// TIA Portal project "Energy_Drink_V15.1" (V15.1) (continued)

       // IF RESET BUTTON OR HMI RESET => RESET RECIPE SELCTION
       IF "Reset_Button" OR "HMI_VAR".Reset_Selection THEN
           "RECIPE_1_DB".Recipe1.Recipe_Act := FALSE;
           "RECIPE_2_DB".Recipe2.Recipe_Act := FALSE;
           "RECIPE_3_DB".Recipe3.Recipe_Act := FALSE;
           "TEST_RECIPE_DB".Test.Recipe_Act := FALSE;
           "Recipe_Num" := 0;
       END_IF;

   END_REGION

   (************************ RECIPE CONFIRMARTION MANAGEMENT **********************************)
   REGION RECIPE SELECTION CONFIRMATION

       // IF ENTER SELECTION IS PRESSED => START PROCESS
       IF "Var_System_DB".System_Generic.Enter_Selection THEN
           "Var_System_DB".System_Generic.Man_Start_Process := true;
       END_IF;

       // IF ENTER SELECTION IS PRESSED => START PROCESS
       IF "HMI_VAR".Enter_Selection THEN
           "HMI_VAR".Start_Process := TRUE;
       END_IF;

   END_REGION
END_FUNCTION

// folder: 05-CONVEYOR MANAGEMENT

FUNCTION "CONVEYOR_BELT" : Void   // FC10, FBD
{ S7_Optimized_Access := 'FALSE' }
VERSION : 0.1
   VAR_INPUT
      Conveyor_Cmd : Bool;
      Time_Act : Time;
   END_VAR
BEGIN

REGION Network 1 (STL): *******************COMMANDS AND CONDITIONS TO MANAGE CONVEYOR BELT********************************************/
   // WHEN SCALE IS FINISHED WEIGHING ALL THE PRODUCTS => BACH IN PROGRESS =1
   // SEND COMMAND TO ACTIVATE THE CONVEYOR BELT
         A     #Conveyor_Cmd;
         FP    "FP_Conveyor_Act";
         S     "Var_System_DB".System_Generic.Mixer_Station;

         A     "Var_System_DB".System_Generic.Mixer_Station;
         FP    "Tag_14";
         =     "Var_System_DB".Conveyor_Belt.Motor_Cmd;


   // TIMER ACTIVATION: IF FN PULSE OF CONVEYOR_CMD => SET TIMER_ACT
         A     #Conveyor_Cmd;
         FN    "FN_Bach_in_Prog";
         =     "Var_System_DB".Conveyor_Belt.Timer_Act;

   // IF TIMER_ACT = 1 => ACTIVATE TIMER
         CALL  TP, "T_CONVEYOR"
         ( IN := "Var_System_DB".Conveyor_Belt.Timer_Act,
           PT := #Time_Act,
           Q  := ,
           ET :=
         );


   // IF TIMER.Q => SEND PULSE TO RESET MOTOR_CMD
         A     "T_CONVEYOR".Q;
         FN    "FN_TIMER.Q";
         R     "Var_System_DB".Conveyor_Belt.M_Stop;


   // SEND PULSE TO SET STOP COMMAND TO ITS NORMAL POSITON "NC" WHEN FN OF FEEDBACK
         A     "Var_System_DB".Conveyor_Belt.M_Feedback;
         FN    "FN_STOP_CMD";
         S     "Var_System_DB".Conveyor_Belt.M_Stop;
         S     "Var_System_DB".System_Generic.Conveyor_Station;


   // RESET CONVEYOR STATION
         A     "AGITATOR_TIMER_DB".Q;
         R     "Var_System_DB".System_Generic.Conveyor_Station;

   // MOTOR MEMORY STATE: IN CASE STOP BUTTON IS PRESSED AND THE  MOTOR WAS ACTIVE,
   // WE WANT TO KEEP THE MOTOR "ON" AFTER THE STOP BUTTON IS REALESED AGAIN
         A     "Var_System_DB".Conveyor_Belt.M_Feedback;
         S     "Var_System_DB".Conveyor_Belt.State;

   // RESET BELT STATE BIT
         AN    "Var_System_DB".System_Generic.Stop_Process;
         AN    "Var_System_DB".System_Generic.System_Failure;
         O(;
         A     "Var_System_DB".System_Generic.Start;
         FN    "Tag_27";
         );
         R     "Var_System_DB".Conveyor_Belt.State;
END_REGION

REGION Network 2: ****************** CONVEYOR BELT MOTOR ACTIVATION********************************************/
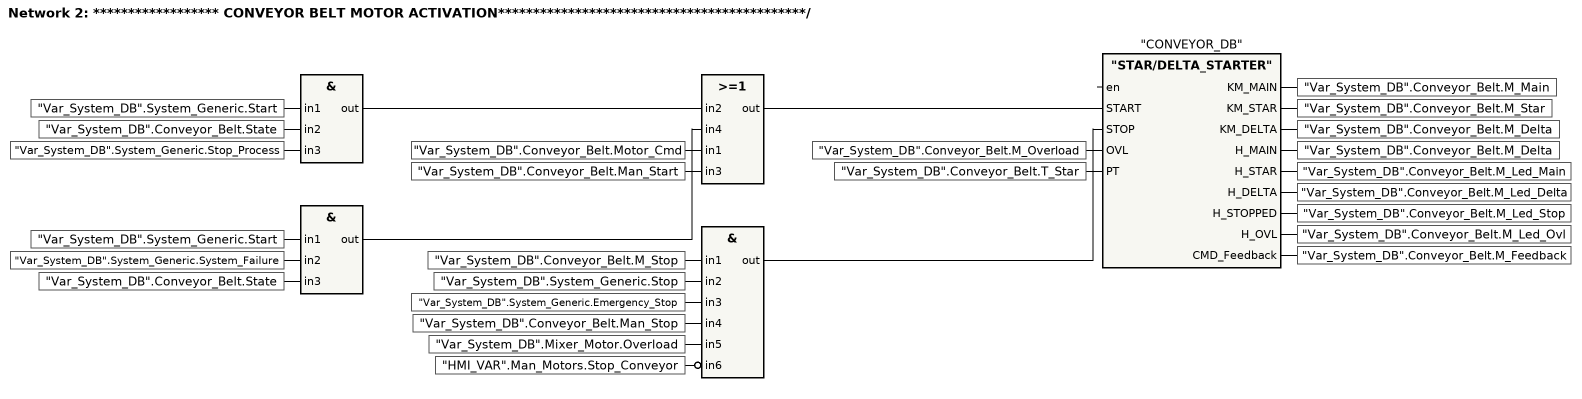
   "CONVEYOR_DB"(START := ("Var_System_DB".System_Generic.Start AND "Var_System_DB".Conveyor_Belt.State AND "Var_System_DB".System_Generic.Stop_Process) OR ("Var_System_DB".System_Generic.Start AND "Var_System_DB".System_Generic.System_Failure AND "Var_System_DB".Conveyor_Belt.State) OR "Var_System_DB".Conveyor_Belt.Motor_Cmd OR "Var_System_DB".Conveyor_Belt.Man_Start,   // "STAR/DELTA_STARTER"
                 STOP := "Var_System_DB".Conveyor_Belt.M_Stop AND "Var_System_DB".System_Generic.Stop AND "Var_System_DB".System_Generic.Emergency_Stop AND "Var_System_DB".Conveyor_Belt.Man_Stop AND "Var_System_DB".Mixer_Motor.Overload AND NOT "HMI_VAR".Man_Motors.Stop_Conveyor,
                 OVL := "Var_System_DB".Conveyor_Belt.M_Overload,
                 PT := "Var_System_DB".Conveyor_Belt.T_Star,
                 KM_MAIN => "Var_System_DB".Conveyor_Belt.M_Main,
                 KM_STAR => "Var_System_DB".Conveyor_Belt.M_Star,
                 KM_DELTA => "Var_System_DB".Conveyor_Belt.M_Delta,
                 H_MAIN => "Var_System_DB".Conveyor_Belt.M_Delta,
                 H_STAR => "Var_System_DB".Conveyor_Belt.M_Led_Main,
                 H_DELTA => "Var_System_DB".Conveyor_Belt.M_Led_Delta,
                 H_STOPPED => "Var_System_DB".Conveyor_Belt.M_Led_Stop,
                 H_OVL => "Var_System_DB".Conveyor_Belt.M_Led_Ovl,
                 CMD_Feedback => "Var_System_DB".Conveyor_Belt.M_Feedback);
END_REGION
END_FUNCTION

// folder: 06-MIXER MANAGEMENT

FUNCTION "MIXER_TANK_MANAGEMENT" : Void   // FC3, FBD
{ S7_Optimized_Access := 'FALSE' }
VERSION : 0.1
BEGIN

REGION Network 1: /***********************MIXER TANK LEVEL*****************************************/
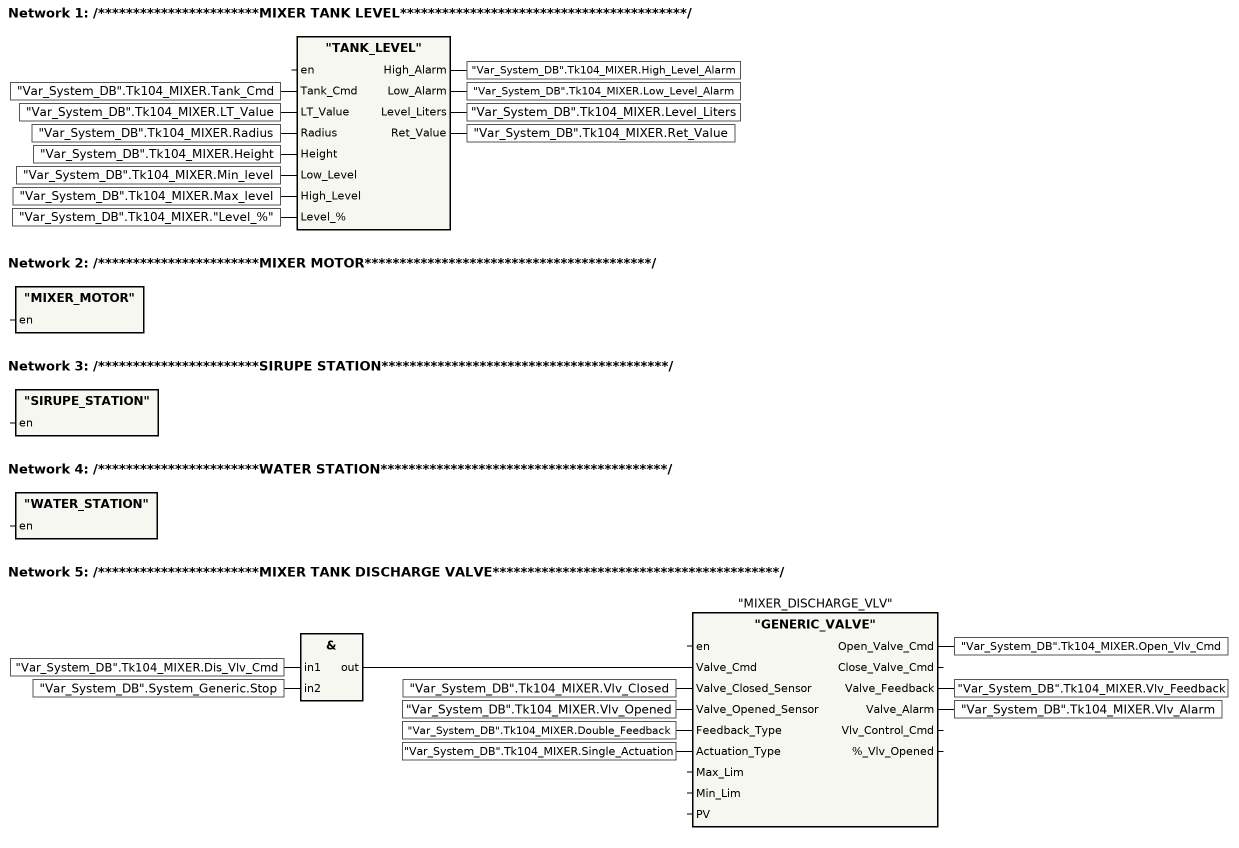
   "TANK_LEVEL"(Tank_Cmd := "Var_System_DB".Tk104_MIXER.Tank_Cmd,
                LT_Value := "Var_System_DB".Tk104_MIXER.LT_Value,
                Radius := "Var_System_DB".Tk104_MIXER.Radius,
                Height := "Var_System_DB".Tk104_MIXER.Height,
                Low_Level := "Var_System_DB".Tk104_MIXER.Min_level,
                High_Level := "Var_System_DB".Tk104_MIXER.Max_level,
                "Level_%" := "Var_System_DB".Tk104_MIXER."Level_%",
                High_Alarm => "Var_System_DB".Tk104_MIXER.High_Level_Alarm,
                Low_Alarm => "Var_System_DB".Tk104_MIXER.Low_Level_Alarm,
                Level_Liters => "Var_System_DB".Tk104_MIXER.Level_Liters,
                Ret_Value => "Var_System_DB".Tk104_MIXER.Ret_Value);
END_REGION

REGION Network 2: /***********************MIXER MOTOR*****************************************/
   "MIXER_MOTOR"();
END_REGION

REGION Network 3: /***********************SIRUPE STATION*****************************************/
   "SIRUPE_STATION"();
END_REGION

REGION Network 4: /***********************WATER STATION*****************************************/
   "WATER_STATION"();
END_REGION

REGION Network 5: /***********************MIXER TANK DISCHARGE VALVE*****************************************/
   "MIXER_DISCHARGE_VLV"(Valve_Cmd := "Var_System_DB".Tk104_MIXER.Dis_Vlv_Cmd AND "Var_System_DB".System_Generic.Stop,   // "GENERIC_VALVE"
                         Valve_Closed_Sensor := "Var_System_DB".Tk104_MIXER.Vlv_Closed,
                         Valve_Opened_Sensor := "Var_System_DB".Tk104_MIXER.Vlv_Opened,
                         Feedback_Type := "Var_System_DB".Tk104_MIXER.Double_Feedback,
                         Actuation_Type := "Var_System_DB".Tk104_MIXER.Single_Actuation,
                         Open_Valve_Cmd => "Var_System_DB".Tk104_MIXER.Open_Vlv_Cmd,
                         Valve_Feedback => "Var_System_DB".Tk104_MIXER.Vlv_Feedback,
                         Valve_Alarm => "Var_System_DB".Tk104_MIXER.Vlv_Alarm);
END_REGION

REGION Network 6 (STL): /***********************TANK CONDITIONS ACTIVATION*****************************************/
   // IF SYSTEM IS ACTIVE AND MIXER STATION => MIXER TANK COMMAND = 1
         A     "Var_System_DB".System_Generic.System_Act;
         A     "Var_System_DB".System_Generic.Mixer_Station;
         =     "Var_System_DB".Tk104_MIXER.Tank_Cmd;

   // IF TANK LEVEL > 15% => SEND COMMAND TO AGITATOR, WATER AND SIRUPE VALVE
         A     "Var_System_DB".Tk104_MIXER.Tank_Cmd;
         A(;
         L     "Var_System_DB".Tk104_MIXER."Level_%";
         L     15;
         >I;
         );
         =     "Var_System_DB".Mixer_Motor.Motor_Cmd;
         =     "Var_System_DB".Sirupe_Valve.Vlv_Cmd;
         =     "Var_System_DB".Water_Valve.Vlv_Cmd;
END_REGION

REGION Network 7 (STL): /***********************TANK CONDITIONS ACTIVATION*****************************************/
   // IF SYSTEM IS ACTIVE, MIXER STATION AND CONVEYOR HAS STOPPED =>
   // ACTIVATE TIMER TO OPEN THE VALVE WHEN ELAPSED TIME IS "ON"
         A     "Var_System_DB".System_Generic.System_Act;
         A     "Var_System_DB".System_Generic.Mixer_Station;
         A     "Var_System_DB".System_Generic.Conveyor_Station;
         FP    "Var_System_DB".Mixer_Motor.FP_Timer;
         =     "Var_System_DB".System_Generic.T_Mixer_Station;

   // TIMER CALL
         CALL  TP, "AGITATOR_TIMER_DB"
         ( IN := "Var_System_DB".System_Generic.T_Mixer_Station,
           PT := T#60S,
           Q  := ,
           ET :=
         );


   // IF FN AGITATOR_TIMER.Q => SEND COMMAND TO ACTIVATE DISCHARGE VALVE
         A     "AGITATOR_TIMER_DB".Q;
         FN    "Var_System_DB".Tk104_MIXER.FN_Agitator;
         S     "Var_System_DB".Tk104_MIXER.Dis_Vlv_Cmd;


   // RESET VALVE COMMAND AND MIXER STATION AND BACH IN PROGRESS
         A     "Var_System_DB".Tk104_MIXER.Dis_Vlv_Cmd;
         A(;
         L     "Var_System_DB".Tk104_MIXER."Level_%";
         L     0;
         ==I;
         );
         R     "Var_System_DB".Tk104_MIXER.Dis_Vlv_Cmd;
         R     "Var_System_DB".System_Generic.Mixer_Station;
         R     "Var_System_DB".System_Generic.Bach_In_Progress;

         ON    "Var_System_DB".System_Generic.System_Act;
         R     "Var_System_DB".Tk104_MIXER.Dis_Vlv_Cmd;
END_REGION
END_FUNCTION

FUNCTION "WATER_STATION" : Void   // FC5, FBD
{ S7_Optimized_Access := 'FALSE' }
VERSION : 0.1
BEGIN

REGION Network 1 (STL): /************************WATER FLOW METER*****************************************/
         CALL  SCALE
         ( IN      := "Var_System_DB".Water_Flow_Meter.Flow_Meter,
           HI_LIM  := "Var_System_DB".Water_Flow_Meter.High_Lim,
           LO_LIM  := "Var_System_DB".Water_Flow_Meter.Low_Lim,
           BIPOLAR := FALSE,
           RET_VAL := "Var_System_DB".Water_Flow_Meter.Ret_Val,
           OUT     := "Var_System_DB".Water_Flow_Meter.Flow_PV
         );
END_REGION

REGION Network 2: /*****************************WATER VALVE***************************************************/
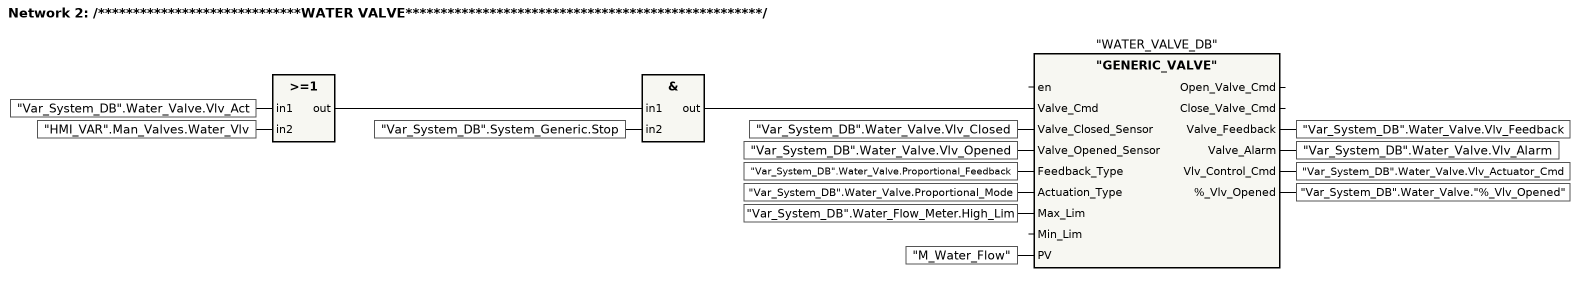
   "WATER_VALVE_DB"(Valve_Cmd := ("Var_System_DB".Water_Valve.Vlv_Act OR "HMI_VAR".Man_Valves.Water_Vlv) AND "Var_System_DB".System_Generic.Stop,   // "GENERIC_VALVE"
                    Valve_Closed_Sensor := "Var_System_DB".Water_Valve.Vlv_Closed,
                    Valve_Opened_Sensor := "Var_System_DB".Water_Valve.Vlv_Opened,
                    Feedback_Type := "Var_System_DB".Water_Valve.Proportional_Feedback,
                    Actuation_Type := "Var_System_DB".Water_Valve.Proportional_Mode,
                    Max_Lim := "Var_System_DB".Water_Flow_Meter.High_Lim,
                    PV := "M_Water_Flow",
                    Valve_Feedback => "Var_System_DB".Water_Valve.Vlv_Feedback,
                    Valve_Alarm => "Var_System_DB".Water_Valve.Vlv_Alarm,
                    Vlv_Control_Cmd => "Var_System_DB".Water_Valve.Vlv_Actuator_Cmd,
                    "%_Vlv_Opened" => "Var_System_DB".Water_Valve."%_Vlv_Opened");
END_REGION

REGION Network 3 (STL)
   // IF VALVE COMMAND SEND PULSE TO ACTIVATE => WATER VALVE
         A     "Var_System_DB".Water_Valve.Vlv_Cmd;
         FP    "Var_System_DB".Water_Valve.FP_Start;
         S     "Var_System_DB".Water_Valve.Vlv_Act;

   // IF MIXWE DISCHARGE VALVE COMMAND SEND PULSE TO DEACTIVATE => WATER VALVE
         A     "Var_System_DB".Tk104_MIXER.Dis_Vlv_Cmd;
         FP    "Var_System_DB".Water_Valve.FP_Stop;
         R     "Var_System_DB".Water_Valve.Vlv_Act;
END_REGION
END_FUNCTION

FUNCTION "SIRUPE_STATION" : Void   // FC7, FBD
{ S7_Optimized_Access := 'FALSE' }
VERSION : 0.1
BEGIN

REGION Network 1 (STL): /************************SIRUPE FLOW METER*****************************************/
         CALL  SCALE
         ( IN      := "Var_System_DB".Sirupe_Flow_Meter.Flow_Meter,
           HI_LIM  := "Var_System_DB".Sirupe_Flow_Meter.Low_Lim,
           LO_LIM  := "Var_System_DB".Sirupe_Flow_Meter.High_Lim,
           BIPOLAR := FALSE,
           RET_VAL := "Var_System_DB".Sirupe_Flow_Meter.Ret_Val,
           OUT     := "Var_System_DB".Sirupe_Flow_Meter.Flow_PV
         );
END_REGION

REGION Network 2 (STL)
         L     "M_Sirupe_Flow";
         L     1000;
         *R;
         T     "Var_System_DB".Sirupe_Valve.Increment_T;
END_REGION

REGION Network 3: /**********************************SIRUPE VALVE*****************************************/
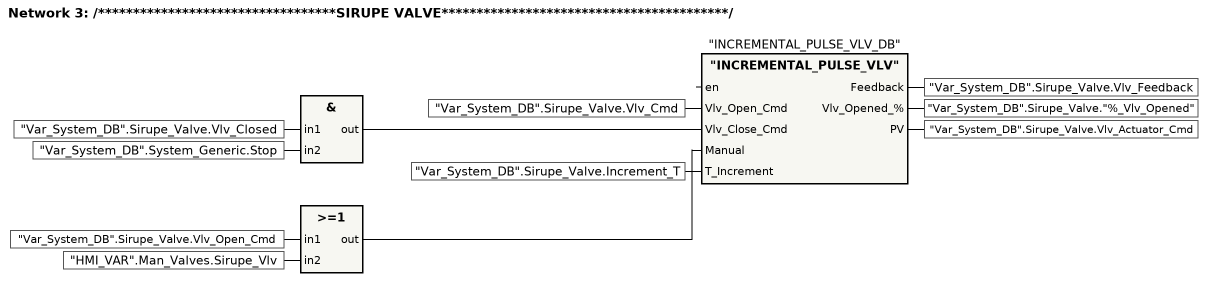
   "INCREMENTAL_PULSE_VLV_DB"(Vlv_Open_Cmd := "Var_System_DB".Sirupe_Valve.Vlv_Cmd,   // "INCREMENTAL_PULSE_VLV"
                           Vlv_Close_Cmd := "Var_System_DB".Sirupe_Valve.Vlv_Closed AND "Var_System_DB".System_Generic.Stop,
                           Manual := "Var_System_DB".Sirupe_Valve.Vlv_Open_Cmd OR "HMI_VAR".Man_Valves.Sirupe_Vlv,
                           T_Increment := "Var_System_DB".Sirupe_Valve.Increment_T,
                           Feedback => "Var_System_DB".Sirupe_Valve.Vlv_Feedback,
                           "Vlv_Opened_%" => "Var_System_DB".Sirupe_Valve."%_Vlv_Opened",
                           PV => "Var_System_DB".Sirupe_Valve.Vlv_Actuator_Cmd);
END_REGION

REGION Network 4 (STL)
   // COMMAND TO CLOSE THE VALVE
         A     "Var_System_DB".Tk104_MIXER.Dis_Vlv_Cmd;
         FP    "Var_System_DB".Sirupe_Valve.FP_Reset;
         =     "Var_System_DB".Sirupe_Valve.Vlv_Closed;
END_REGION
END_FUNCTION

FUNCTION "MIXER_MOTOR" : Void   // FC13, FBD
{ S7_Optimized_Access := 'FALSE' }
VERSION : 0.1
BEGIN

REGION Network 1 (STL): *******************COMMANDS AND CONDITIONS TO MANAGE AGITATOR********************************************/
   // IF MOTOR CMD FP => SEND COMMAND TO ACTIVATE AGITATOR
         A     "Var_System_DB".Mixer_Motor.Motor_Cmd;
         FP    "Var_System_DB".Mixer_Motor.FP_Start;
         O     "Var_System_DB".Mixer_Motor.Man_Start;
         =     "Var_System_DB".Mixer_Motor.Cmd_Start;

   // IF MOTOR CMD FN => SEND COMMAND TO DEACTIVATE AGITATOR
         A     "Var_System_DB".Mixer_Motor.Motor_Cmd;
         FN    "Var_System_DB".Mixer_Motor.FN_Stop;
         ON    "Var_System_DB".Mixer_Motor.Man_Stop;
         R     "Var_System_DB".Mixer_Motor.Cmd_Stop;


   // IF CMD STOP NOT ACTIVE AND MOTOR PV = 0 => SET BACK CMD STOP = 1
         AN    "Var_System_DB".Mixer_Motor.Cmd_Stop;
         A(;
         L     "Var_System_DB".Mixer_Motor.PV;
         L     0;
         ==I;
         );
         S     "Var_System_DB".Mixer_Motor.Cmd_Stop;


   // RESET MIXER MOTOR STATE:
   // IF NOT STOP PROCESS AND NOT SYSTEM FAILURE (NOT OVERLOAD) AND MOTOR_PV == 0
   // OR NEGATIVE EDGE OF GENERIC START
         AN    "Var_System_DB".System_Generic.Stop_Process;
         AN    "Var_System_DB".System_Generic.System_Failure;
         A(;
         L     "Var_System_DB".Mixer_Motor.PV;
         L     0;
         ==I;
         );
         O(;
         A     "Var_System_DB".System_Generic.Start;
         FN    "Tag_26";
         );
         R     "Var_System_DB".Mixer_Motor.State;


   // MOTOR MEMORY STATE IN CASE STOP BUTTON PRESSED AND THE  MOTOR WAS ACTIVE
   // WE WANT TO KEEP THE MOTOR ON AFTER THE STOP BUTTON
         A     "Var_System_DB".Mixer_Motor.Feedback;
         S     "Var_System_DB".Mixer_Motor.State;
END_REGION

REGION Network 2
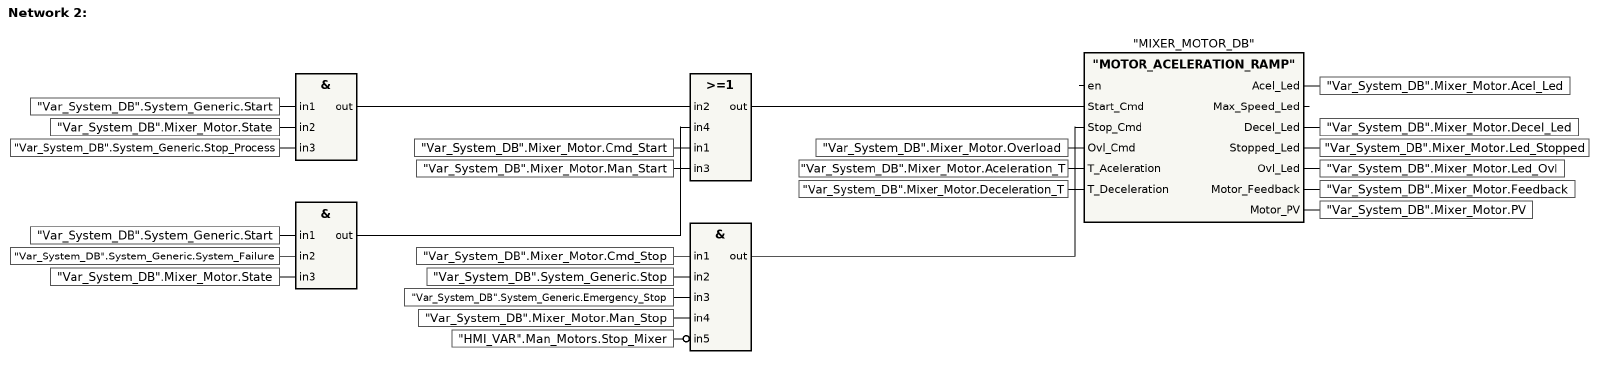
   "MIXER_MOTOR_DB"(Start_Cmd := ("Var_System_DB".System_Generic.Start AND "Var_System_DB".Mixer_Motor.State AND "Var_System_DB".System_Generic.Stop_Process) OR ("Var_System_DB".System_Generic.Start AND "Var_System_DB".System_Generic.System_Failure AND "Var_System_DB".Mixer_Motor.State) OR "Var_System_DB".Mixer_Motor.Cmd_Start OR "Var_System_DB".Mixer_Motor.Man_Start,   // "MOTOR_ACELERATION_RAMP"
                    Stop_Cmd := "Var_System_DB".Mixer_Motor.Cmd_Stop AND "Var_System_DB".System_Generic.Stop AND "Var_System_DB".System_Generic.Emergency_Stop AND "Var_System_DB".Mixer_Motor.Man_Stop AND NOT "HMI_VAR".Man_Motors.Stop_Mixer,
                    Ovl_Cmd := "Var_System_DB".Mixer_Motor.Overload,
                    T_Aceleration := "Var_System_DB".Mixer_Motor.Aceleration_T,
                    T_Deceleration := "Var_System_DB".Mixer_Motor.Deceleration_T,
                    Acel_Led => "Var_System_DB".Mixer_Motor.Acel_Led,
                    Decel_Led => "Var_System_DB".Mixer_Motor.Decel_Led,
                    Stopped_Led => "Var_System_DB".Mixer_Motor.Led_Stopped,
                    Ovl_Led => "Var_System_DB".Mixer_Motor.Led_Ovl,
                    Motor_Feedback => "Var_System_DB".Mixer_Motor.Feedback,
                    Motor_PV => "Var_System_DB".Mixer_Motor.PV);
END_REGION
END_FUNCTION

// folder: FBs

FUNCTION_BLOCK "GENERIC_VALVE"   // FB1, SCL
{ S7_Optimized_Access := 'FALSE' }
VERSION : 0.1
   VAR_INPUT
      Valve_Cmd : Bool;   // Enable valve command
      Valve_Closed_Sensor : Bool;   // Valve closed position
      Valve_Opened_Sensor : Bool;   // Valve opened position
      Feedback_Type : Int;   // "0" = No feedback / "1"= Single disFeedback / "2"= Single EnFeedback / "3" = Double Feedback / "4" = Proportional
      Actuation_Type : Int;
      Max_Lim : Real;
      Min_Lim : Real;
      PV : Real;
   END_VAR
   VAR_OUTPUT
      Open_Valve_Cmd : Bool;
      Close_Valve_Cmd : Bool;
      Valve_Feedback : Bool;   // "1" If the valve is open, "0" otherwise
      Valve_Alarm : Bool;
      Vlv_Control_Cmd : Int;
      "%_Vlv_Opened" : DInt;
   END_VAR
   VAR
      M_Vlv_Closed : Bool;
      M_Vlv_Opened : Bool;
      Ret_Vlv : Word;
   END_VAR
   VAR_TEMP
      Temp_Process_Signal : Real;
   END_VAR
   VAR CONSTANT
      No_Feedback : Int := 0;
      Single_En_Feedback : Int := 1;
      Single_Dis_Feedback : Int := 2;
      Double_Feedback : Int := 3;
      Proportional_Feedback : Int := 4;
      Single_Actuation : Int := 1;
      Double_Actuation : Int := 2;
      Proportional_Mode : Int := 3;
      Inverse_Mode : Int := 4;
      Control_Loop : Int := 5;
   END_VAR
BEGIN
   (*
   *File: FB GENERIC VALVE 
   * Author: Jaime Calvente Mieres
   * Date: 18-05-2022
   * Description: This FB will be used to control a valve. Depending on 
     the users input, the valve could act as Single actuation,
     Double actuation or Proportional mode.
   *)



   (*This Case Statement will be used to map the process sensors to
   the internal variables used for the program logic, based on the
   Feedback Type or (Type of Valve) used in each process.*)
   REGION FEEDBACK_TYPE

       CASE #Feedback_Type OF

           #No_Feedback:
               ;

           #Single_En_Feedback:
               #M_Vlv_Opened := #Valve_Opened_Sensor;

           #Single_Dis_Feedback:
               #M_Vlv_Closed := #Valve_Closed_Sensor;

           #Double_Feedback:
               #M_Vlv_Closed := #Valve_Closed_Sensor;
               #M_Vlv_Opened := #Valve_Opened_Sensor;

           #Proportional_Feedback:
               #M_Vlv_Closed := #Valve_Closed_Sensor;
               #M_Vlv_Opened := #Valve_Opened_Sensor;

           ELSE  // Statement section ELSE
               ;
       END_CASE;


   END_REGION


   // IF VALVE COMMAND ACTIVE
   IF #Valve_Cmd THEN

   (*This Case Statement will be used to Set the type of Actuation will be used
   depending on the types of Valves the process has.*)
       REGION ACTUATION_TYPE

           CASE #Actuation_Type OF

                   // SINGLE ACTUATION VALVES    
               #Single_Actuation:

                   IF #Valve_Closed_Sensor THEN
                       #Open_Valve_Cmd := true;
                   END_IF;

                   // DOUBLE ACTUATION VALVES        
               #Double_Actuation:

                   IF #M_Vlv_Closed THEN
                       #Open_Valve_Cmd := true;
                   ELSIF #M_Vlv_Opened THEN
                       #Open_Valve_Cmd := false;
                   END_IF;

                   (*
                       PROPORTIONAL ACTUATION VALVES 
                   *)

                   // PROPORTIONAL MODE
               #Proportional_Mode:
                   #Temp_Process_Signal := #PV;
                   #Ret_Vlv := UNSCALE(IN := #Temp_Process_Signal, HI_LIM := #Max_Lim, LO_LIM := #Min_Lim, BIPOLAR := false, OUT => #Vlv_Control_Cmd);
                   #"%_Vlv_Opened" := ROUND((#Vlv_Control_Cmd * 100.0) / 27648);

                   // INVERSE MODE
               #Inverse_Mode:
                   #Temp_Process_Signal := #PV;
                   #Ret_Vlv := UNSCALE(IN := #Temp_Process_Signal, HI_LIM := #Min_Lim, LO_LIM := #Max_Lim, BIPOLAR := false, OUT => #Vlv_Control_Cmd);
                   #"%_Vlv_Opened" := ROUND((#Vlv_Control_Cmd * 100.0) / 27648);

                   // PID CONTROL MODE
               #Control_Loop:
                   #Temp_Process_Signal := #PV;
                   #Ret_Vlv := UNSCALE(IN := #Temp_Process_Signal, HI_LIM := #Max_Lim, LO_LIM := #Min_Lim, BIPOLAR := false, OUT => #Vlv_Control_Cmd);
                   #"%_Vlv_Opened" := ROUND((#Vlv_Control_Cmd * 100.0) / 27648);

           END_CASE;

       END_REGION




   // IF NOT VALVE COMMAND
   ELSE
       // KEEP THE VALVE IN A CLOSED POSITION.
       #Open_Valve_Cmd := false;
       #Close_Valve_Cmd := true;

       // IF VALVE ALREARY CLOSED  => SET COMMAND TO "0"
       IF #M_Vlv_Closed THEN
           #Close_Valve_Cmd := false;
       END_IF;

       // IF PROPORTIONAL MODES ACTIVE =>VALVE RETURN "0" 
       #Vlv_Control_Cmd := 0;
       #"%_Vlv_Opened" := 0;
   END_IF;
END_FUNCTION_BLOCK

FUNCTION_BLOCK "STAR/DELTA_STARTER"   // FB2, STL
{ S7_Optimized_Access := 'FALSE' }
VERSION : 0.1
// STAR-DELTA GENERIC STARTER
   VAR_INPUT
      START : Bool;   // START ACTION
      STOP : Bool;   // STOP ACTION
      OVL : Bool;   // MOTOR OVERLOAD
      PT : Time;
   END_VAR
   VAR_OUTPUT
      KM_MAIN : Bool;   // MAIN CONTACTOR
      KM_STAR : Bool;   // STAR CONTACTOR
      KM_DELTA : Bool;   // DELTA CONTACTOR
      H_MAIN : Bool;   // MAIN LED
      H_STAR : Bool;   // STAR LED
      H_DELTA : Bool;   // DELTA LED
      H_STOPPED : Bool;   // STOP LED
      H_OVL : Bool;   // OVERLOAD LED
      CMD_Feedback : Bool;
   END_VAR
   VAR
      SYSTEM_OK : Bool;
      M_MAIN : Bool;   // VAR MEMORY MAIN CONTACTOR
      M_STAR : Bool;   // VAR MEMORY STAR CONTACTOR
      M_DELTA : Bool;   // VAR MEMORY DELTA CONTACTOR
      M_TIMER : Bool;   // VAR MEMORY TIMER
      "TIME" : Time;
      STAR_TIMER : TON;
   END_VAR
   // STAR_TIMER.PT := T#0MS;
BEGIN

REGION Network 1: ***************************** SYSTEM MANAGEMENT ********************************************/ / SYSTEM STATUS
   // WHILE OVL AND STOP = 1, SYSTEM OK
         A     #OVL;
         A     #STOP;
         =     #SYSTEM_OK;
END_REGION

REGION Network 2: ***************************** STAR MODE CONDITIONS ********************************************/ / VAR MEMORY TIMER AND STAR CONTACTOR ACTIVATION
   // SET MEMORY TO ACTIVATE TIMER AND STAR CONTACTOR CONDITION
         A     #SYSTEM_OK;
         AN    #STAR_TIMER.Q;
         A(;
         A     #START;
         O     #M_STAR;
         );
         S     #M_TIMER;
         =     #M_STAR;

   // IF TIME.Q = TRUE, RESET M_TIMER
         A     #STAR_TIMER.Q;
         R     #M_TIMER;

   // IF S_TIMER = TRUE, ACTIVATE TIMER
         CALL  #STAR_TIMER
         ( IN := #M_TIMER,
           PT := #PT,
           Q  := ,
           ET := #STAR_TIMER.ET
         );
END_REGION

REGION Network 3: ***************************** STAR KM AND LED ACTIVATION ********************************************/ / STAR CONTACTOR
   // WHILE M_STAR = 1, STAR CONTACTOR AND LED ARE "ON"
         A     #M_STAR;
         =     #KM_STAR;
         =     #H_STAR;
END_REGION

REGION Network 4: ***************************** MAIN KM ACTIVATION CONDITIONS ********************************************/ / VAR MEMORY MAIN CONTACTOR
   // CONDITIONS TO ACTIVATE M_MAIN CONTACTOR
         A     #SYSTEM_OK;
         A(;
         A     #M_STAR;
         O     #M_MAIN;
         );
         =     #M_MAIN;

   // WHILE M_MAIN = 1, MAIN CONTACTOR AND LED ARE "ON"
         A     #M_MAIN;
         =     #KM_MAIN;
         =     #H_MAIN;
END_REGION

REGION Network 5: ***************************** DELTA KM ACTIVATION CONDITIONS ********************************************/ / VAR MEMORY DELTA CONTACTOR
   // CONDITIONS TO ACTIVATE M_DELTA CONTACTOR
         A     #SYSTEM_OK;
         A     #M_MAIN;
         AN    #M_STAR;
         =     #M_DELTA;

   // WHILE M_DELTA = 1, DELTA CONTACTOR AND LED ARE "ON"
         A     #M_DELTA;
         =     #KM_DELTA;
         =     #H_DELTA;
         =     #CMD_Feedback;
END_REGION

REGION Network 6: *****************************STOP LED ACTIVATION ********************************************/ / STOP LED
         AN    #STOP;
         ON    #M_MAIN;
         =     #H_STOPPED;
END_REGION

REGION Network 7: *****************************OVERLOAD LED ACTIVATION ********************************************/ / OVERLOAD LED
         AN    #OVL;
         =     #H_OVL;
END_REGION
END_FUNCTION_BLOCK

FUNCTION_BLOCK "MOTOR_ACELERATION_RAMP"   // FB3, STL
{ S7_Optimized_Access := 'FALSE' }
VERSION : 0.1
   VAR_INPUT
      Start_Cmd : Bool;
      Stop_Cmd : Bool;
      Ovl_Cmd : Bool;
   END_VAR
   VAR_OUTPUT
      Acel_Led : Bool;
      Max_Speed_Led : Bool;
      Decel_Led : Bool;
      Stopped_Led : Bool;
      Ovl_Led : Bool;
      Motor_Feedback : Bool;
      Motor_PV : Int;
   END_VAR
   VAR_IN_OUT
      T_Aceleration : Time;
      T_Deceleration : Time;
   END_VAR
   VAR
      Aceleration_State : Bool;
      Deceleration_State : Bool;
      Full_load : Bool;
      FP_Stop : Bool;
      Ret_Val_Acel : Word;
      Ret_Val_Decel : Word;
      Motor_Cmd : Int;
      Aceleration : Real;
      Deceleration : Real;
      Max_Lim : Real;
      Low_Lim : Real := 0.0;
      Aceleration_Timer : TP;
      Deceleration_Timer : TP;
   END_VAR
BEGIN

REGION Network 1: SI PULSAMOS MARCHA Y NO ESTA DECELERANDO => ACTIVAMOS ACELERACION / /************************** ACELERATION MODE *****************************************/
   // CONDITIONS TO SET ACELEREATION STATE
         A     #Ovl_Cmd;
         A     #Start_Cmd;
         AN    #Deceleration_State;
         R     #Deceleration_State;
         S     #Aceleration_State;

   // RESET CONDITIONS ACELERATION STATE
         A(;
         L     #Motor_Cmd;
         L     27648;
         ==I;
         );
         R     #Aceleration_State;

   // IF ACELERATION STATE IS ACTIVE => SEND COMMAND TO GRADUALLY INCREASE MOTOR VELOCITY
         A     #Aceleration_State;
         JCN   _100;

   // ANOLOG SIGNAL UNSCALING TO GENEREATE THE ACELERATION BASED ON A TIMER

         CALL  UNSCALE
         ( IN      := #Aceleration,
           HI_LIM  := #Max_Lim,
           LO_LIM  := #Low_Lim,
           BIPOLAR := FALSE,
           RET_VAL := #Ret_Val_Acel,
           OUT     := #Motor_Cmd
         );

   // SETTING THE MAX LIMIT
         L     #T_Aceleration;
         DTR;
         T     #Max_Lim;

   // MAPPING VAR FOR CONSULTING
         L     #Motor_Cmd;
         T     #Motor_PV;
   _100: NOP   0;


   // TIMER TO GENERATE THE ACELERETAION VARIABLE
         CALL  #Aceleration_Timer
         ( IN := #Aceleration_State,
           PT := #T_Aceleration,
           Q  := ,
           ET := #Aceleration_Timer.ET
         );

   // CONVERTIN THE ELAPSED TIME INTO REAL => TO ASIGN AS INPUT OF THE AO ACELERATION
         L     #Aceleration_Timer.ET;
         DTR;
         T     #Aceleration;
END_REGION

REGION Network 2: SI PULSAMOS PARO Y NO ESTÁ ACELERANDO => RAMPA DECELERACION ACTIVA / /************************** DECELERATION MODE *****************************************/
   // CONDITIONS TO SET THE DECELERATION STATE
         AN    #Stop_Cmd;
         FP    #FP_Stop;  // IT IS AN FP DUE TO THE FACT THAT IS "NC"
         AN    #Aceleration_State;
         A(;
         L     #Motor_Cmd;
         L     0;
         <>I;
         );
         S     #Deceleration_State;

   // IF DECELERATION STATE IS ACTIVE => SEND COMMAND TO GRADUALLY DECREASE MOTOR SPEED
         A     #Deceleration_State;
         JCN   _105;

   // ANOLOG SIGNAL UNSCALING TO GENEREATE THE DECELERATION BASED ON A TIMER

         CALL  UNSCALE
         ( IN      := #Deceleration,
           HI_LIM  := #Low_Lim,
           LO_LIM  := #Max_Lim,
           BIPOLAR := FALSE,
           RET_VAL := #Ret_Val_Decel,
           OUT     := #Motor_Cmd
         );

   // MAPPING VAR FOR CONSULTING
         L     #Motor_Cmd;
         T     #Motor_PV;

   // SETTING THE MAX LIMIT
         L     #T_Deceleration;
         DTR;
         T     #Max_Lim;

   _105: NOP   0;


   // TIMER TO GENERATE THE DECELERETAION VARIABLE
         CALL  #Deceleration_Timer
         ( IN := #Deceleration_State,
           PT := #T_Deceleration,
           Q  := ,
           ET := #Deceleration_Timer.ET
         );


   // CONVERTIN THE ELAPSED TIME INTO REAL => TO ASIGN AS INPUT OF THE AO DECELERATION
         L     #Deceleration_Timer.ET;
         DTR;
         T     #Deceleration;
END_REGION

REGION Network 3: CONDITIONS FOR EMERGENCY STOP BY OVERLOAD OR STOP BUTTON WHILE ACELERATING / /******************************STOPPING MODE *****************************************/
   // IF MOTOR OVERLOAD OR STOP BUTTON AND ACELERATION => EMERGENCY STOP
         AN    #Ovl_Cmd;
         O(;
         AN    #Stop_Cmd;
         A     #Aceleration_State;
         );
         JCN   _108;
         L     0;
         T     #Motor_PV;
         T     #Motor_Cmd;

   _108: NOP   0;
END_REGION

REGION Network 4: ACELERATION AND MAX SPEED LED ACTIVATION / /******************************LED ACTIVATIONS *****************************************/
   // LED START ACTIVATION
         A     #Aceleration_State;
         A(;
         L     #Motor_Cmd;
         L     27648;
         <I;
         );
         A(;
         L     #Motor_Cmd;
         L     0;
         >I;
         );
         =     #Acel_Led;  // ACELERATION LED ACTIVE


   // LED MAX SPEED ACTIVATION
         A(;
         L     #Motor_Cmd;
         L     27648;
         ==I;
         );
         =     #Full_load;
         =     #Max_Speed_Led;  // MAX SPEED LED ACTIVE

   // DECELERATION LED ACTIVATION
         A     #Deceleration_State;
         A(;
         L     #Motor_Cmd;
         L     27648;
         <I;
         );
         A(;
         L     #Motor_Cmd;
         L     0;
         >I;
         );
         =     #Decel_Led;

   // STOPPED LED ACTIVATION
         A(;
         L     #Motor_Cmd;
         L     0;
         ==I;
         );
         R     #Deceleration_State;

   // STOPPED LED DEACTIVATION
         A     #Stop_Cmd;
         AN    #Aceleration_State;
         AN    #Full_load;
         S     #Stopped_Led;

         A     #Start_Cmd;
         R     #Stopped_Led;

   // OVERLOAD LED ACTIVATION
         AN    #Ovl_Cmd;
         =     #Ovl_Led;
END_REGION

REGION Network 5: *******************MOTOR FEEDBACK********************************************/
   // CONDITIONS FOR MOTOR FEEDBACK
         A     #Aceleration_State;
         O     #Full_load;
         =     #Motor_Feedback;
END_REGION
END_FUNCTION_BLOCK

FUNCTION_BLOCK "INCREMENTAL_PULSE_VLV"   // FB4, STL
{ S7_Optimized_Access := 'FALSE' }
VERSION : 0.1
   VAR_INPUT
      Vlv_Open_Cmd : Bool;
      Vlv_Close_Cmd : Bool;
      Manual : Bool;
   END_VAR
   VAR_OUTPUT
      Feedback : Bool;
      "Vlv_Opened_%" : DInt;
      PV : Int;
   END_VAR
   VAR_IN_OUT
      T_Increment : Time;
   END_VAR
   VAR
      Incremental_State : Bool;
      Pulse_Loop : Bool;
      FP_Start : Bool;
      FP_Stop : Bool;
      Ret_Val_Acel : Word;
      Valve_Cmd : Int;
      Increment : Real;
      Max_Lim : Real;
      Low_Lim : Real;
      Incremental_Timer : TP;
   END_VAR
BEGIN

REGION Network 1: SI PULSAMOS MARCHA Y NO ESTA DECELERANDO => ACTIVAMOS ACELERACION / /******************************PULSE INCREMENTAL MODE *****************************************/
   // PULSAR MARCHA PARA ACTIVAR EL MOTOR CON RAMPA DE ACELERACION
         A     #Vlv_Open_Cmd;
         FP    #FP_Start;
         S     #Incremental_State;

   // RESET CONDITIONS ACELERATION STATE
         A     #Incremental_State;
         A(;
         L     #Valve_Cmd;
         L     27648;
         ==I;
         );
         JCN   INCR2;
         L     0;
         T     #Increment;
         T     #Valve_Cmd;
         T     #PV;
   INCR2:NOP   0;

